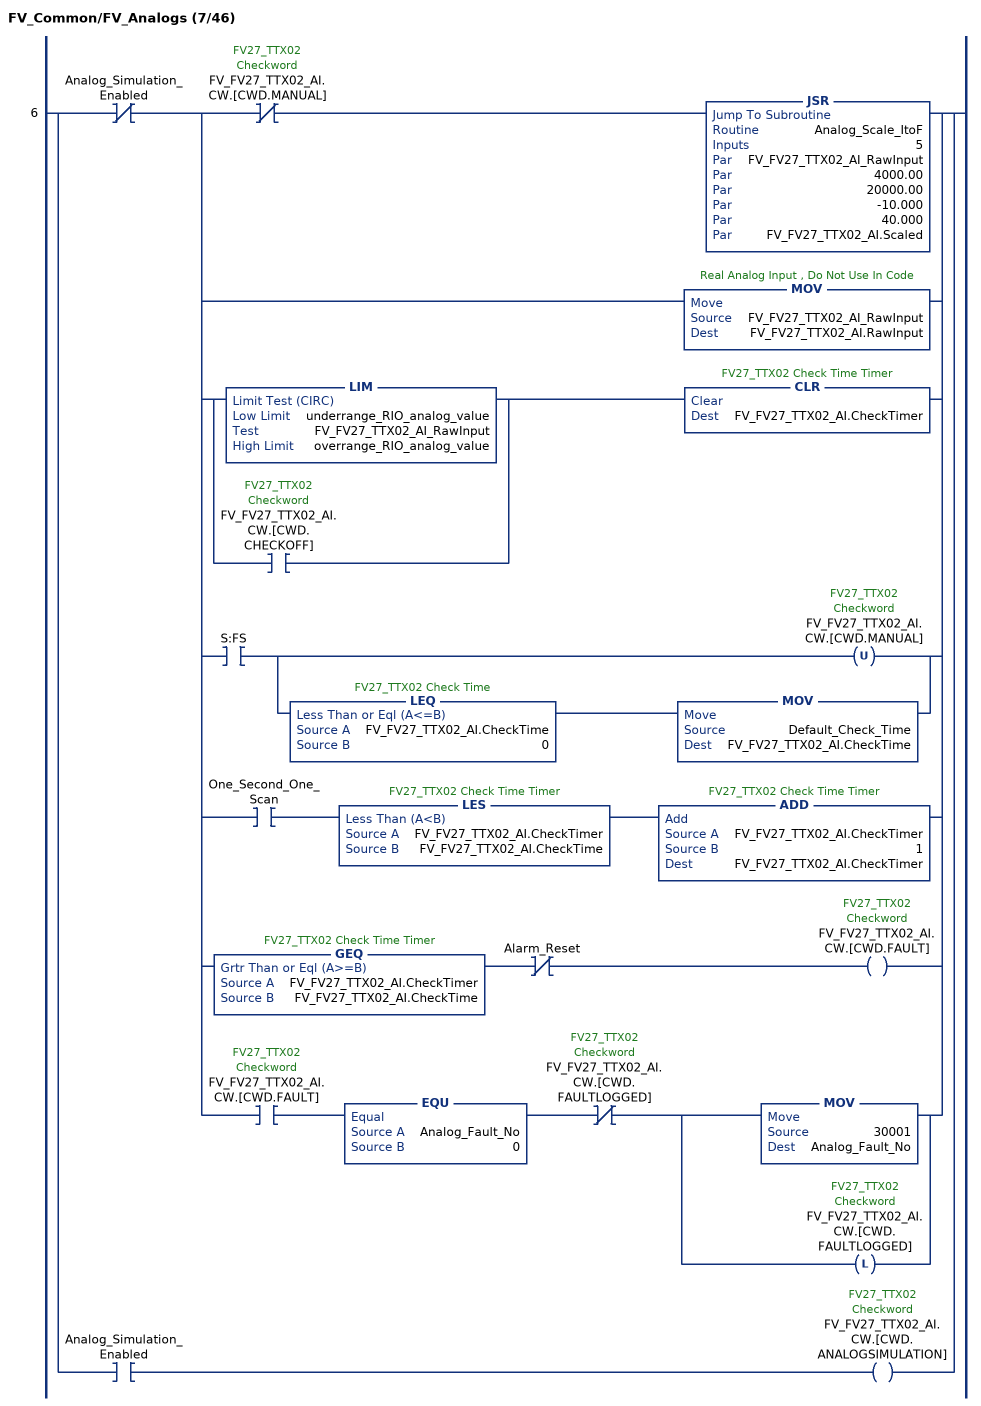
   6: [XIO(Analog_Simulation_Enabled) [XIO(FV_FV27_TTX02_AI.CW.[CWD.MANUAL]) JSR(Analog_Scale_ItoF,5,FV_FV27_TTX02_AI_RawInput,4000.00,20000.00,-10.000,40.000,FV_FV27_TTX02_AI.Scaled) ,MOV(FV_FV27_TTX02_AI_RawInput,FV_FV27_TTX02_AI.RawInput) ,[LIM(underrange_RIO_analog_value,FV_FV27_TTX02_AI_RawInput,overrange_RIO_analog_value) ,XIC(FV_FV27_TTX02_AI.CW.[CWD.CHECKOFF]) ] CLR(FV_FV27_TTX02_AI.CheckTimer) ,XIC(S:FS) [OTU(FV_FV27_TTX02_AI.CW.[CWD.MANUAL]) ,LEQ(FV_FV27_TTX02_AI.CheckTime,0) MOV(Default_Check_Time,FV_FV27_TTX02_AI.CheckTime) ] ,XIC(One_Second_One_Scan) LES(FV_FV27_TTX02_AI.CheckTimer,FV_FV27_TTX02_AI.CheckTime) ADD(FV_FV27_TTX02_AI.CheckTimer,1,FV_FV27_TTX02_AI.CheckTimer) ,GEQ(FV_FV27_TTX02_AI.CheckTimer,FV_FV27_TTX02_AI.CheckTime) XIO(Alarm_Reset) OTE(FV_FV27_TTX02_AI.CW.[CWD.FAULT]) ,XIC(FV_FV27_TTX02_AI.CW.[CWD.FAULT]) EQU(Analog_Fault_No,0) XIO(FV_FV27_TTX02_AI.CW.[CWD.FAULTLOGGED]) [MOV(30001,Analog_Fault_No) ,OTL(FV_FV27_TTX02_AI.CW.[CWD.FAULTLOGGED]) ] ] ,XIC(Analog_Simulation_Enabled) OTE(FV_FV27_TTX02_AI.CW.[CWD.ANALOGSIMULATION]) ];
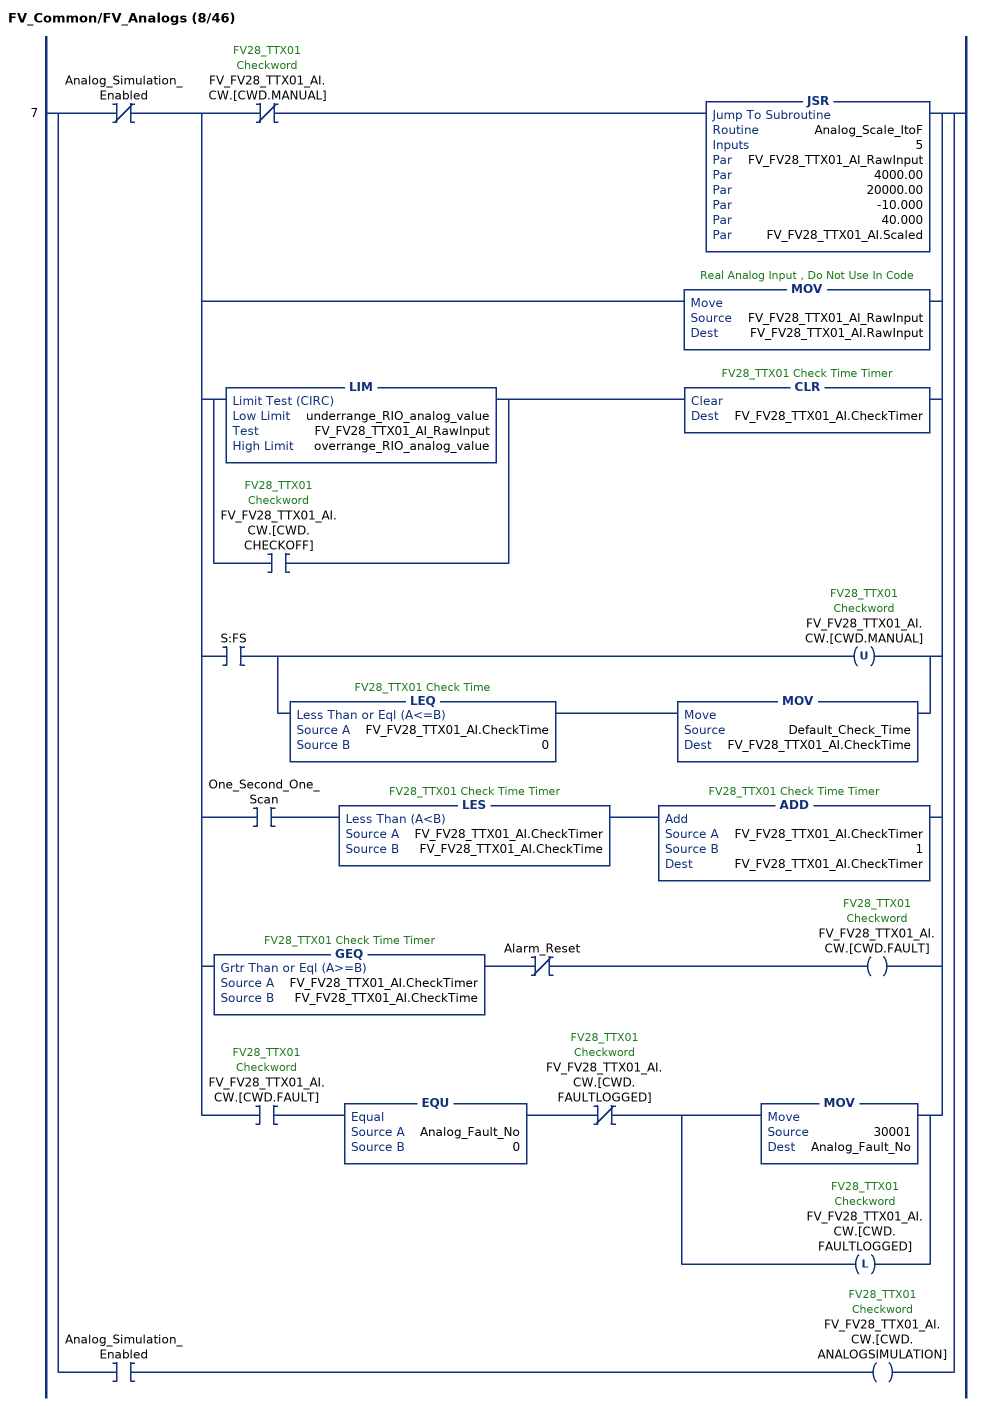
   7: [XIO(Analog_Simulation_Enabled) [XIO(FV_FV28_TTX01_AI.CW.[CWD.MANUAL]) JSR(Analog_Scale_ItoF,5,FV_FV28_TTX01_AI_RawInput,4000.00,20000.00,-10.000,40.000,FV_FV28_TTX01_AI.Scaled) ,MOV(FV_FV28_TTX01_AI_RawInput,FV_FV28_TTX01_AI.RawInput) ,[LIM(underrange_RIO_analog_value,FV_FV28_TTX01_AI_RawInput,overrange_RIO_analog_value) ,XIC(FV_FV28_TTX01_AI.CW.[CWD.CHECKOFF]) ] CLR(FV_FV28_TTX01_AI.CheckTimer) ,XIC(S:FS) [OTU(FV_FV28_TTX01_AI.CW.[CWD.MANUAL]) ,LEQ(FV_FV28_TTX01_AI.CheckTime,0) MOV(Default_Check_Time,FV_FV28_TTX01_AI.CheckTime) ] ,XIC(One_Second_One_Scan) LES(FV_FV28_TTX01_AI.CheckTimer,FV_FV28_TTX01_AI.CheckTime) ADD(FV_FV28_TTX01_AI.CheckTimer,1,FV_FV28_TTX01_AI.CheckTimer) ,GEQ(FV_FV28_TTX01_AI.CheckTimer,FV_FV28_TTX01_AI.CheckTime) XIO(Alarm_Reset) OTE(FV_FV28_TTX01_AI.CW.[CWD.FAULT]) ,XIC(FV_FV28_TTX01_AI.CW.[CWD.FAULT]) EQU(Analog_Fault_No,0) XIO(FV_FV28_TTX01_AI.CW.[CWD.FAULTLOGGED]) [MOV(30001,Analog_Fault_No) ,OTL(FV_FV28_TTX01_AI.CW.[CWD.FAULTLOGGED]) ] ] ,XIC(Analog_Simulation_Enabled) OTE(FV_FV28_TTX01_AI.CW.[CWD.ANALOGSIMULATION]) ];
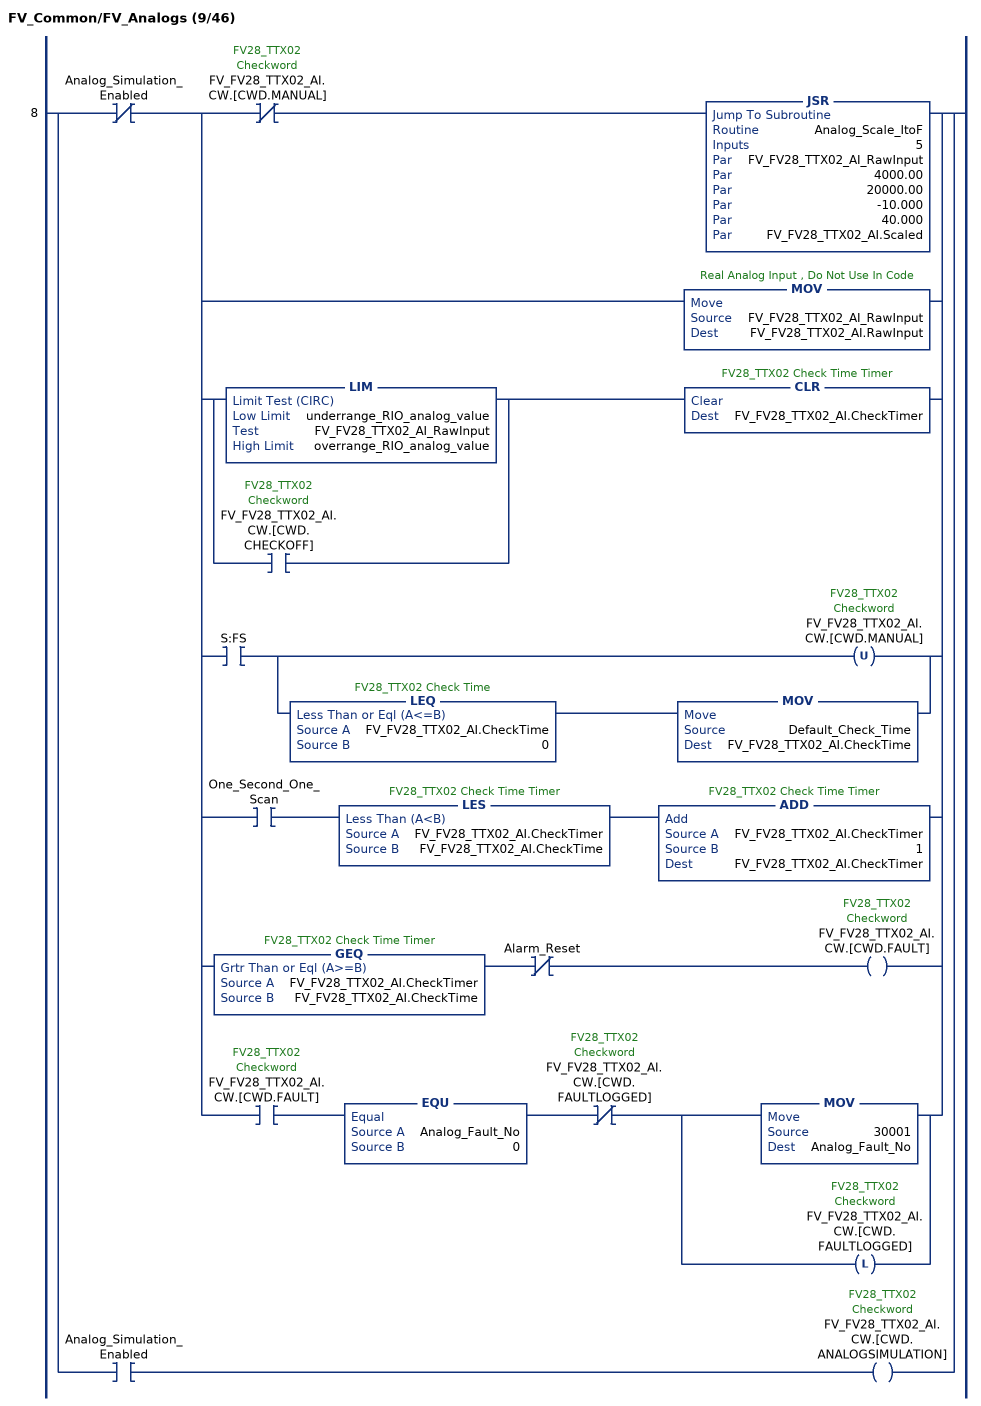
   8: [XIO(Analog_Simulation_Enabled) [XIO(FV_FV28_TTX02_AI.CW.[CWD.MANUAL]) JSR(Analog_Scale_ItoF,5,FV_FV28_TTX02_AI_RawInput,4000.00,20000.00,-10.000,40.000,FV_FV28_TTX02_AI.Scaled) ,MOV(FV_FV28_TTX02_AI_RawInput,FV_FV28_TTX02_AI.RawInput) ,[LIM(underrange_RIO_analog_value,FV_FV28_TTX02_AI_RawInput,overrange_RIO_analog_value) ,XIC(FV_FV28_TTX02_AI.CW.[CWD.CHECKOFF]) ] CLR(FV_FV28_TTX02_AI.CheckTimer) ,XIC(S:FS) [OTU(FV_FV28_TTX02_AI.CW.[CWD.MANUAL]) ,LEQ(FV_FV28_TTX02_AI.CheckTime,0) MOV(Default_Check_Time,FV_FV28_TTX02_AI.CheckTime) ] ,XIC(One_Second_One_Scan) LES(FV_FV28_TTX02_AI.CheckTimer,FV_FV28_TTX02_AI.CheckTime) ADD(FV_FV28_TTX02_AI.CheckTimer,1,FV_FV28_TTX02_AI.CheckTimer) ,GEQ(FV_FV28_TTX02_AI.CheckTimer,FV_FV28_TTX02_AI.CheckTime) XIO(Alarm_Reset) OTE(FV_FV28_TTX02_AI.CW.[CWD.FAULT]) ,XIC(FV_FV28_TTX02_AI.CW.[CWD.FAULT]) EQU(Analog_Fault_No,0) XIO(FV_FV28_TTX02_AI.CW.[CWD.FAULTLOGGED]) [MOV(30001,Analog_Fault_No) ,OTL(FV_FV28_TTX02_AI.CW.[CWD.FAULTLOGGED]) ] ] ,XIC(Analog_Simulation_Enabled) OTE(FV_FV28_TTX02_AI.CW.[CWD.ANALOGSIMULATION]) ];
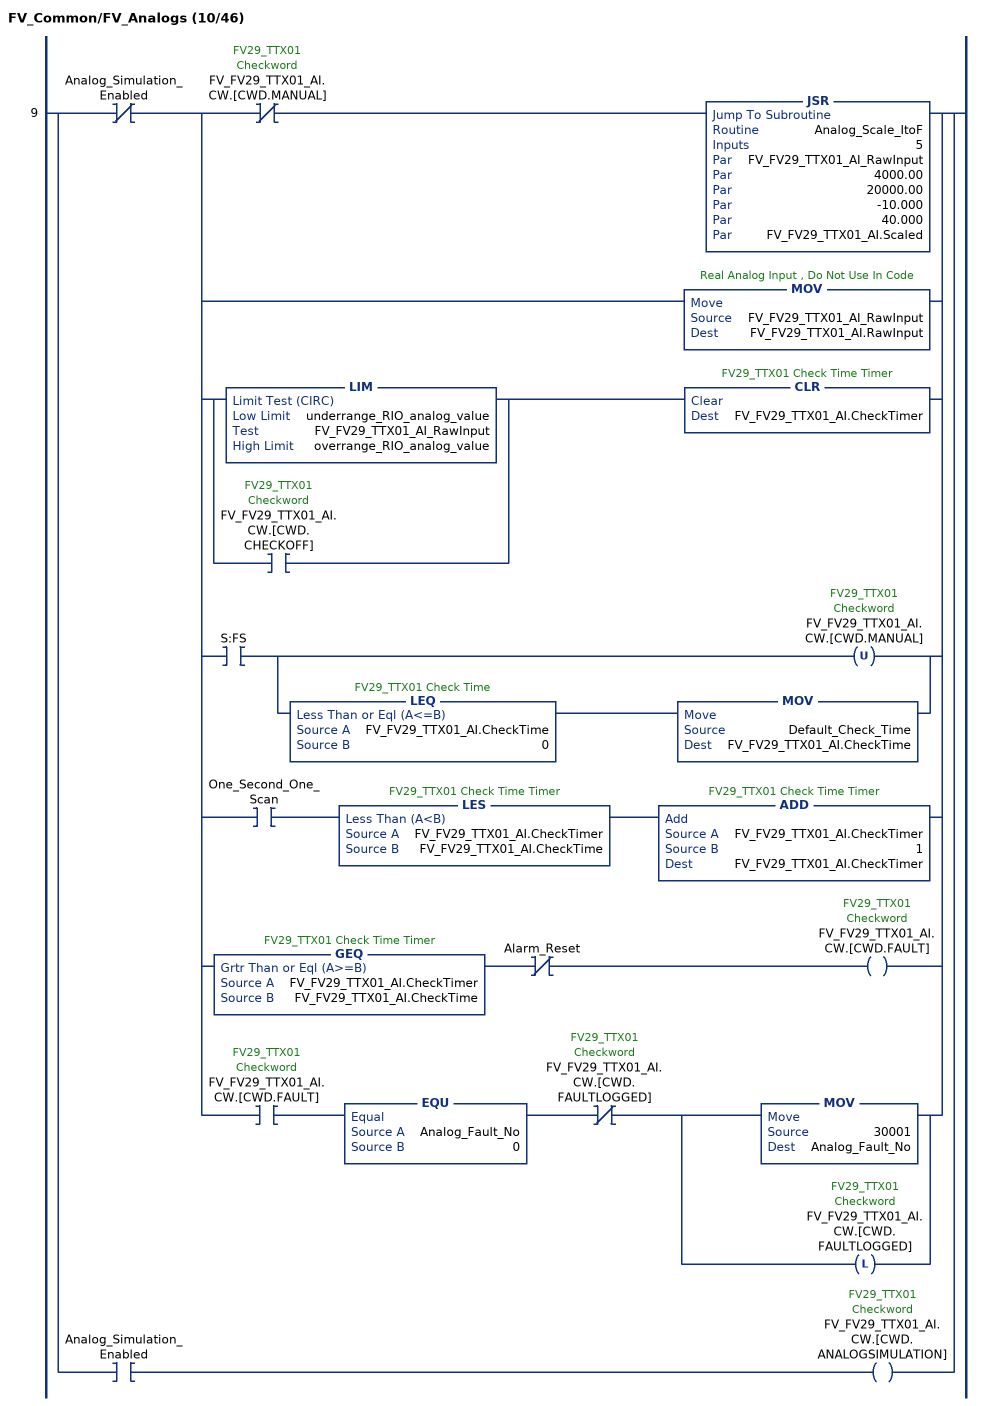
   9: [XIO(Analog_Simulation_Enabled) [XIO(FV_FV29_TTX01_AI.CW.[CWD.MANUAL]) JSR(Analog_Scale_ItoF,5,FV_FV29_TTX01_AI_RawInput,4000.00,20000.00,-10.000,40.000,FV_FV29_TTX01_AI.Scaled) ,MOV(FV_FV29_TTX01_AI_RawInput,FV_FV29_TTX01_AI.RawInput) ,[LIM(underrange_RIO_analog_value,FV_FV29_TTX01_AI_RawInput,overrange_RIO_analog_value) ,XIC(FV_FV29_TTX01_AI.CW.[CWD.CHECKOFF]) ] CLR(FV_FV29_TTX01_AI.CheckTimer) ,XIC(S:FS) [OTU(FV_FV29_TTX01_AI.CW.[CWD.MANUAL]) ,LEQ(FV_FV29_TTX01_AI.CheckTime,0) MOV(Default_Check_Time,FV_FV29_TTX01_AI.CheckTime) ] ,XIC(One_Second_One_Scan) LES(FV_FV29_TTX01_AI.CheckTimer,FV_FV29_TTX01_AI.CheckTime) ADD(FV_FV29_TTX01_AI.CheckTimer,1,FV_FV29_TTX01_AI.CheckTimer) ,GEQ(FV_FV29_TTX01_AI.CheckTimer,FV_FV29_TTX01_AI.CheckTime) XIO(Alarm_Reset) OTE(FV_FV29_TTX01_AI.CW.[CWD.FAULT]) ,XIC(FV_FV29_TTX01_AI.CW.[CWD.FAULT]) EQU(Analog_Fault_No,0) XIO(FV_FV29_TTX01_AI.CW.[CWD.FAULTLOGGED]) [MOV(30001,Analog_Fault_No) ,OTL(FV_FV29_TTX01_AI.CW.[CWD.FAULTLOGGED]) ] ] ,XIC(Analog_Simulation_Enabled) OTE(FV_FV29_TTX01_AI.CW.[CWD.ANALOGSIMULATION]) ];
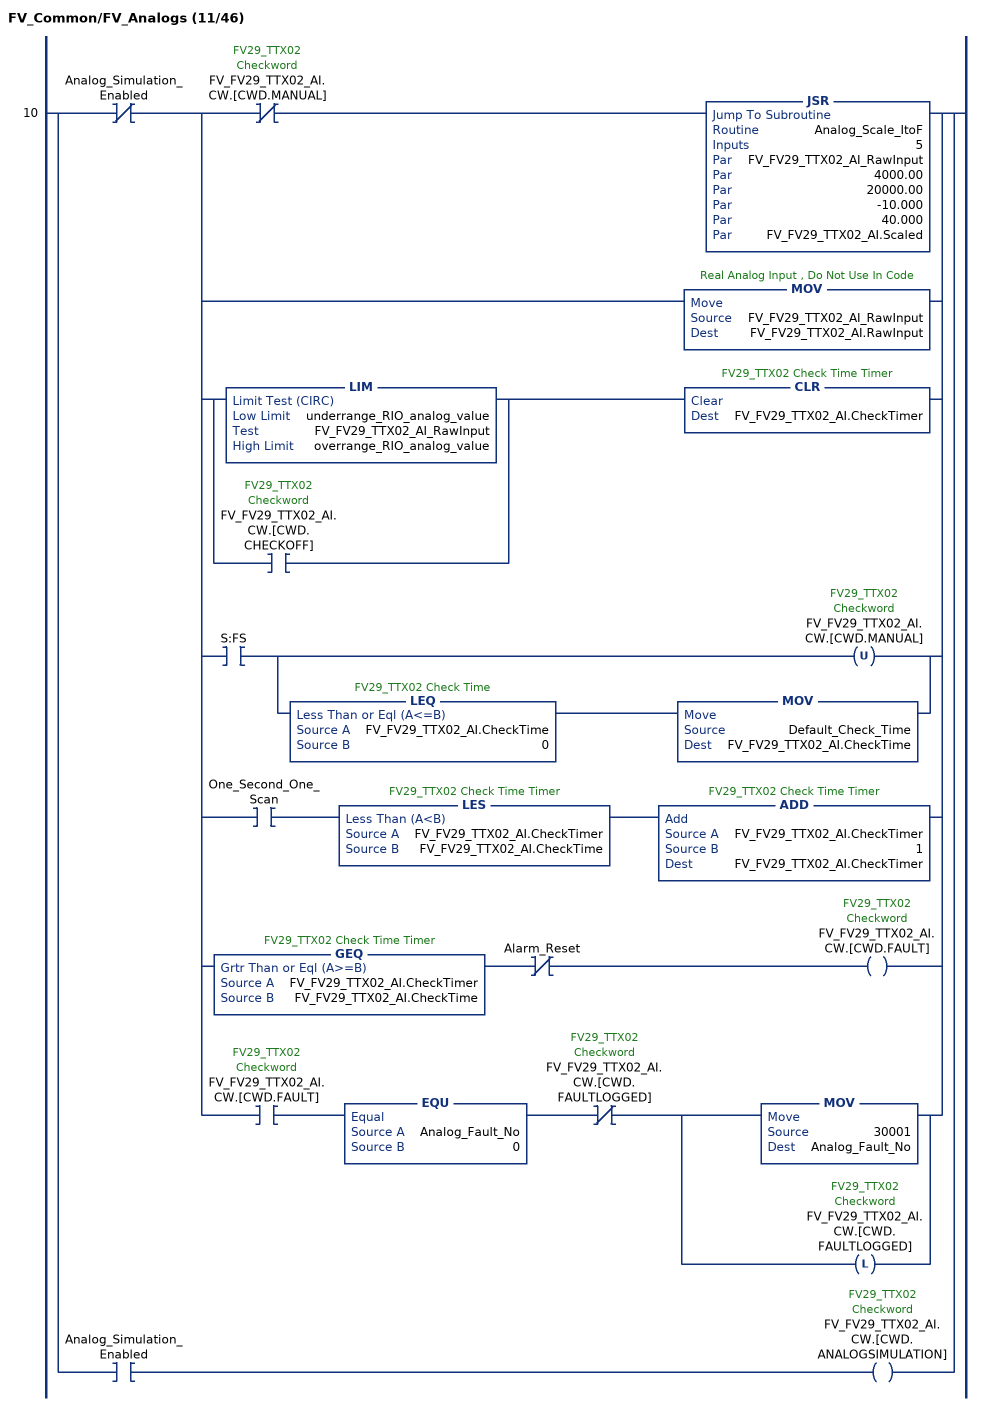
   10: [XIO(Analog_Simulation_Enabled) [XIO(FV_FV29_TTX02_AI.CW.[CWD.MANUAL]) JSR(Analog_Scale_ItoF,5,FV_FV29_TTX02_AI_RawInput,4000.00,20000.00,-10.000,40.000,FV_FV29_TTX02_AI.Scaled) ,MOV(FV_FV29_TTX02_AI_RawInput,FV_FV29_TTX02_AI.RawInput) ,[LIM(underrange_RIO_analog_value,FV_FV29_TTX02_AI_RawInput,overrange_RIO_analog_value) ,XIC(FV_FV29_TTX02_AI.CW.[CWD.CHECKOFF]) ] CLR(FV_FV29_TTX02_AI.CheckTimer) ,XIC(S:FS) [OTU(FV_FV29_TTX02_AI.CW.[CWD.MANUAL]) ,LEQ(FV_FV29_TTX02_AI.CheckTime,0) MOV(Default_Check_Time,FV_FV29_TTX02_AI.CheckTime) ] ,XIC(One_Second_One_Scan) LES(FV_FV29_TTX02_AI.CheckTimer,FV_FV29_TTX02_AI.CheckTime) ADD(FV_FV29_TTX02_AI.CheckTimer,1,FV_FV29_TTX02_AI.CheckTimer) ,GEQ(FV_FV29_TTX02_AI.CheckTimer,FV_FV29_TTX02_AI.CheckTime) XIO(Alarm_Reset) OTE(FV_FV29_TTX02_AI.CW.[CWD.FAULT]) ,XIC(FV_FV29_TTX02_AI.CW.[CWD.FAULT]) EQU(Analog_Fault_No,0) XIO(FV_FV29_TTX02_AI.CW.[CWD.FAULTLOGGED]) [MOV(30001,Analog_Fault_No) ,OTL(FV_FV29_TTX02_AI.CW.[CWD.FAULTLOGGED]) ] ] ,XIC(Analog_Simulation_Enabled) OTE(FV_FV29_TTX02_AI.CW.[CWD.ANALOGSIMULATION]) ];
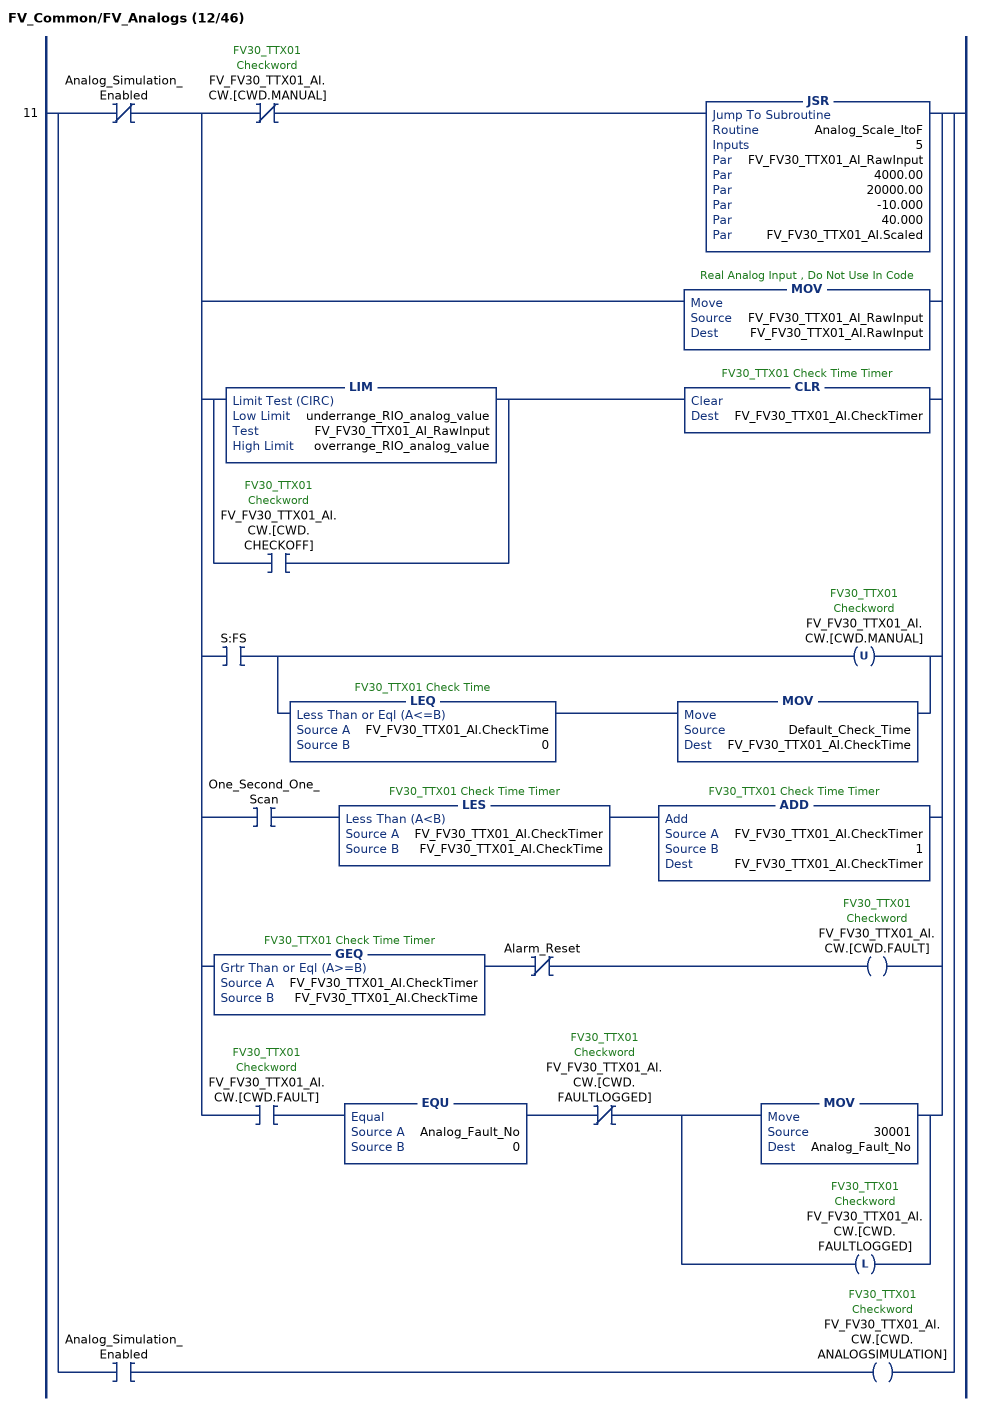
   11: [XIO(Analog_Simulation_Enabled) [XIO(FV_FV30_TTX01_AI.CW.[CWD.MANUAL]) JSR(Analog_Scale_ItoF,5,FV_FV30_TTX01_AI_RawInput,4000.00,20000.00,-10.000,40.000,FV_FV30_TTX01_AI.Scaled) ,MOV(FV_FV30_TTX01_AI_RawInput,FV_FV30_TTX01_AI.RawInput) ,[LIM(underrange_RIO_analog_value,FV_FV30_TTX01_AI_RawInput,overrange_RIO_analog_value) ,XIC(FV_FV30_TTX01_AI.CW.[CWD.CHECKOFF]) ] CLR(FV_FV30_TTX01_AI.CheckTimer) ,XIC(S:FS) [OTU(FV_FV30_TTX01_AI.CW.[CWD.MANUAL]) ,LEQ(FV_FV30_TTX01_AI.CheckTime,0) MOV(Default_Check_Time,FV_FV30_TTX01_AI.CheckTime) ] ,XIC(One_Second_One_Scan) LES(FV_FV30_TTX01_AI.CheckTimer,FV_FV30_TTX01_AI.CheckTime) ADD(FV_FV30_TTX01_AI.CheckTimer,1,FV_FV30_TTX01_AI.CheckTimer) ,GEQ(FV_FV30_TTX01_AI.CheckTimer,FV_FV30_TTX01_AI.CheckTime) XIO(Alarm_Reset) OTE(FV_FV30_TTX01_AI.CW.[CWD.FAULT]) ,XIC(FV_FV30_TTX01_AI.CW.[CWD.FAULT]) EQU(Analog_Fault_No,0) XIO(FV_FV30_TTX01_AI.CW.[CWD.FAULTLOGGED]) [MOV(30001,Analog_Fault_No) ,OTL(FV_FV30_TTX01_AI.CW.[CWD.FAULTLOGGED]) ] ] ,XIC(Analog_Simulation_Enabled) OTE(FV_FV30_TTX01_AI.CW.[CWD.ANALOGSIMULATION]) ];
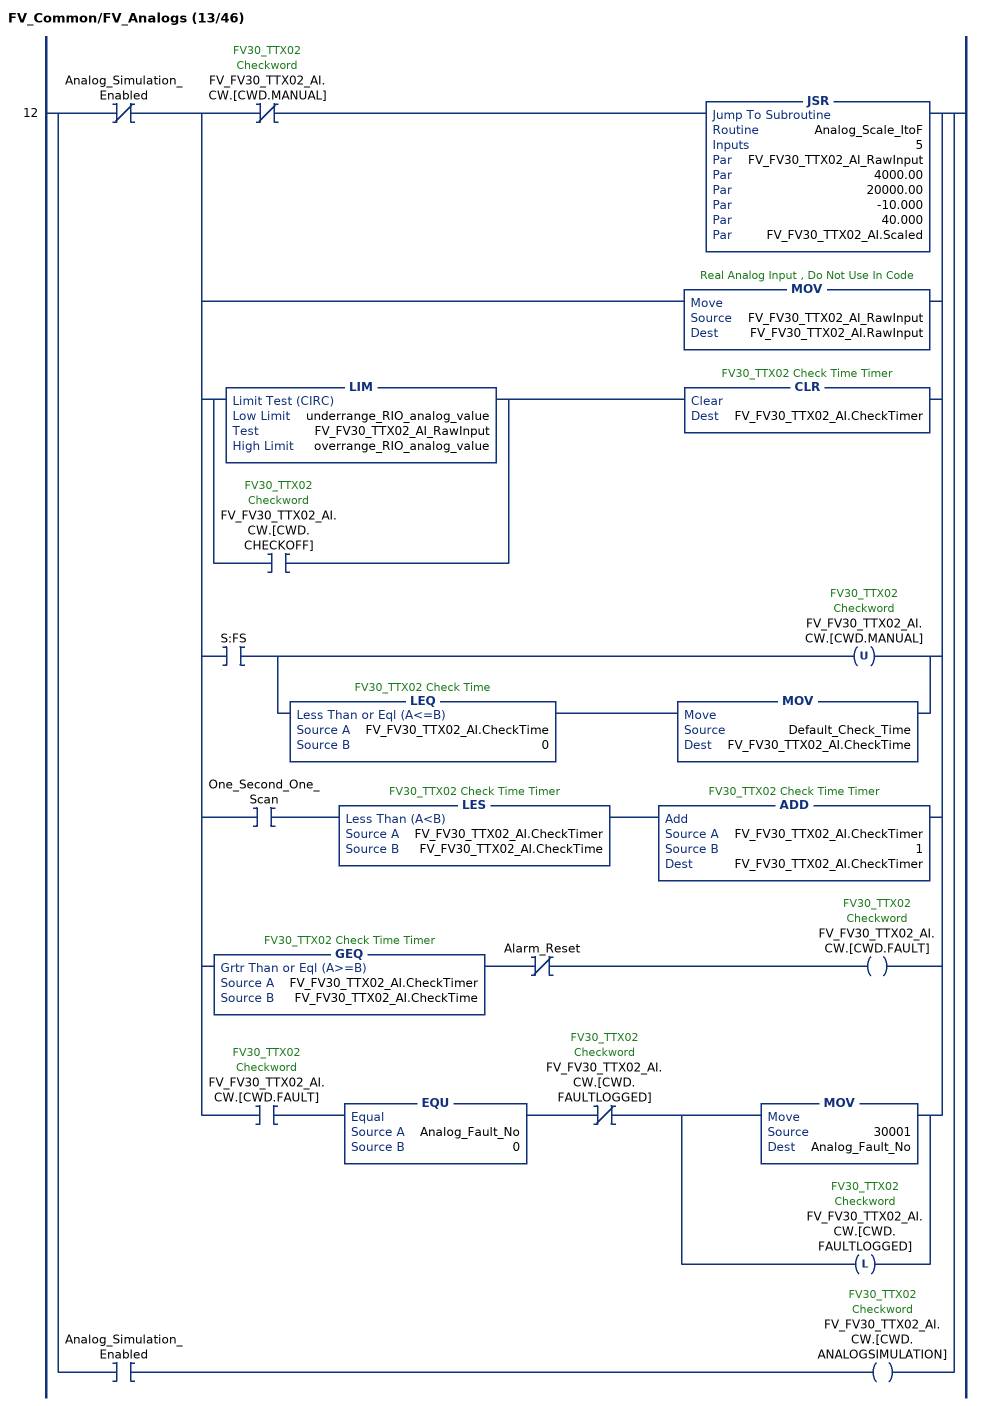
   12: [XIO(Analog_Simulation_Enabled) [XIO(FV_FV30_TTX02_AI.CW.[CWD.MANUAL]) JSR(Analog_Scale_ItoF,5,FV_FV30_TTX02_AI_RawInput,4000.00,20000.00,-10.000,40.000,FV_FV30_TTX02_AI.Scaled) ,MOV(FV_FV30_TTX02_AI_RawInput,FV_FV30_TTX02_AI.RawInput) ,[LIM(underrange_RIO_analog_value,FV_FV30_TTX02_AI_RawInput,overrange_RIO_analog_value) ,XIC(FV_FV30_TTX02_AI.CW.[CWD.CHECKOFF]) ] CLR(FV_FV30_TTX02_AI.CheckTimer) ,XIC(S:FS) [OTU(FV_FV30_TTX02_AI.CW.[CWD.MANUAL]) ,LEQ(FV_FV30_TTX02_AI.CheckTime,0) MOV(Default_Check_Time,FV_FV30_TTX02_AI.CheckTime) ] ,XIC(One_Second_One_Scan) LES(FV_FV30_TTX02_AI.CheckTimer,FV_FV30_TTX02_AI.CheckTime) ADD(FV_FV30_TTX02_AI.CheckTimer,1,FV_FV30_TTX02_AI.CheckTimer) ,GEQ(FV_FV30_TTX02_AI.CheckTimer,FV_FV30_TTX02_AI.CheckTime) XIO(Alarm_Reset) OTE(FV_FV30_TTX02_AI.CW.[CWD.FAULT]) ,XIC(FV_FV30_TTX02_AI.CW.[CWD.FAULT]) EQU(Analog_Fault_No,0) XIO(FV_FV30_TTX02_AI.CW.[CWD.FAULTLOGGED]) [MOV(30001,Analog_Fault_No) ,OTL(FV_FV30_TTX02_AI.CW.[CWD.FAULTLOGGED]) ] ] ,XIC(Analog_Simulation_Enabled) OTE(FV_FV30_TTX02_AI.CW.[CWD.ANALOGSIMULATION]) ];
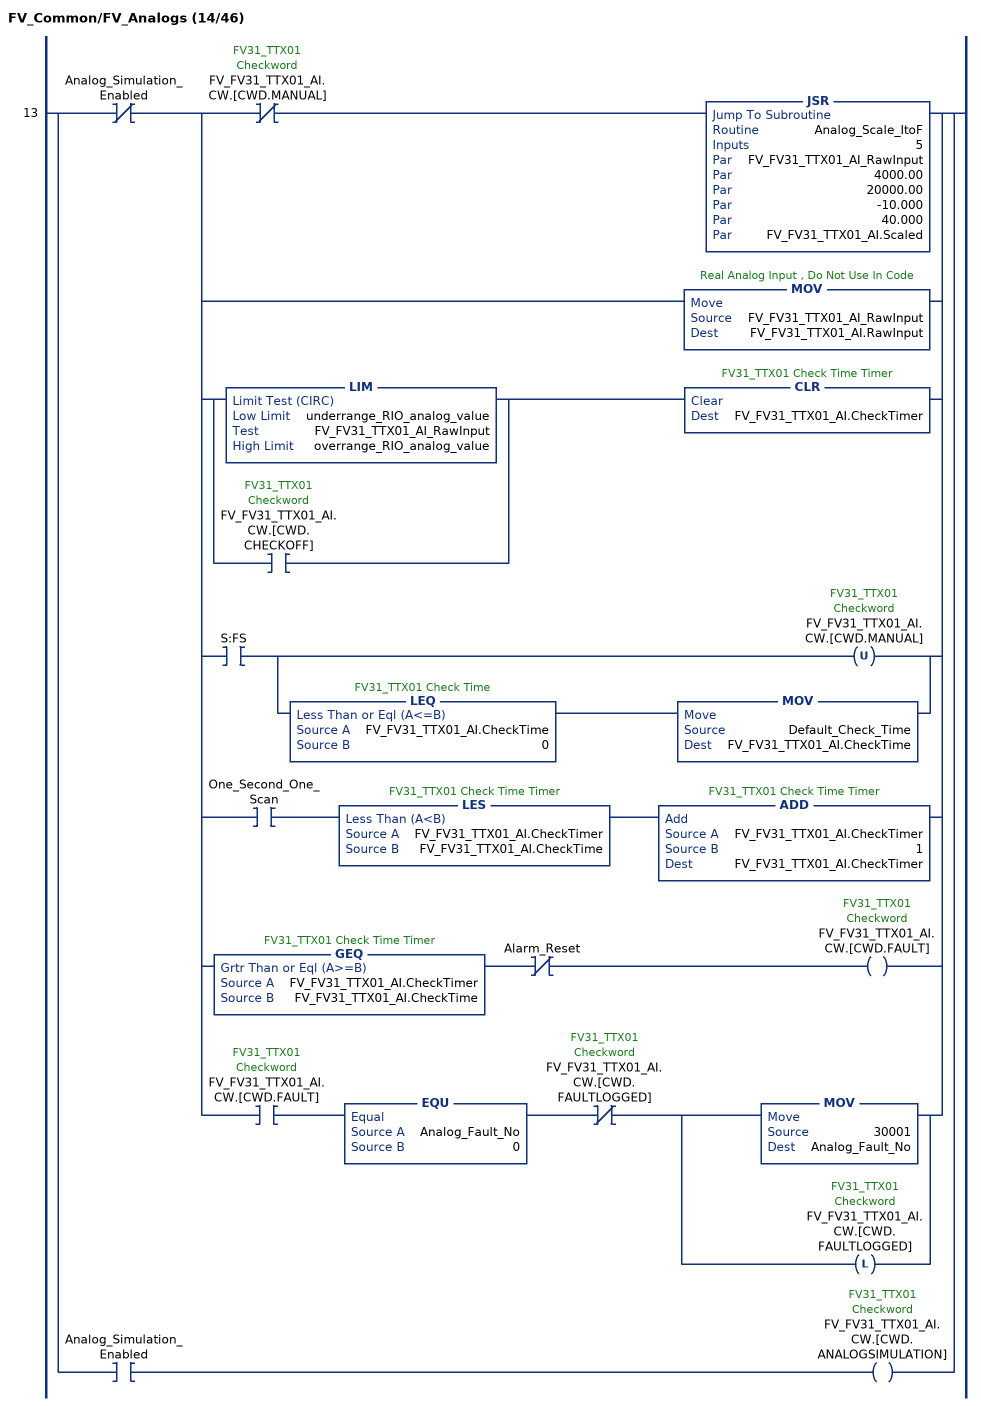
   13: [XIO(Analog_Simulation_Enabled) [XIO(FV_FV31_TTX01_AI.CW.[CWD.MANUAL]) JSR(Analog_Scale_ItoF,5,FV_FV31_TTX01_AI_RawInput,4000.00,20000.00,-10.000,40.000,FV_FV31_TTX01_AI.Scaled) ,MOV(FV_FV31_TTX01_AI_RawInput,FV_FV31_TTX01_AI.RawInput) ,[LIM(underrange_RIO_analog_value,FV_FV31_TTX01_AI_RawInput,overrange_RIO_analog_value) ,XIC(FV_FV31_TTX01_AI.CW.[CWD.CHECKOFF]) ] CLR(FV_FV31_TTX01_AI.CheckTimer) ,XIC(S:FS) [OTU(FV_FV31_TTX01_AI.CW.[CWD.MANUAL]) ,LEQ(FV_FV31_TTX01_AI.CheckTime,0) MOV(Default_Check_Time,FV_FV31_TTX01_AI.CheckTime) ] ,XIC(One_Second_One_Scan) LES(FV_FV31_TTX01_AI.CheckTimer,FV_FV31_TTX01_AI.CheckTime) ADD(FV_FV31_TTX01_AI.CheckTimer,1,FV_FV31_TTX01_AI.CheckTimer) ,GEQ(FV_FV31_TTX01_AI.CheckTimer,FV_FV31_TTX01_AI.CheckTime) XIO(Alarm_Reset) OTE(FV_FV31_TTX01_AI.CW.[CWD.FAULT]) ,XIC(FV_FV31_TTX01_AI.CW.[CWD.FAULT]) EQU(Analog_Fault_No,0) XIO(FV_FV31_TTX01_AI.CW.[CWD.FAULTLOGGED]) [MOV(30001,Analog_Fault_No) ,OTL(FV_FV31_TTX01_AI.CW.[CWD.FAULTLOGGED]) ] ] ,XIC(Analog_Simulation_Enabled) OTE(FV_FV31_TTX01_AI.CW.[CWD.ANALOGSIMULATION]) ];